   // IF ACELERATION STATE IS ACTIVE => SEND COMMAND TO GRADUALLY INCREASE MOTOR VELOCITY
         A     #Incremental_State;
         JCN   _100;

   // ANOLOG SIGNAL UNSCALING TO GENEREATE THE INCREMENTAL ACTION BASED ON A TIMER

         CALL  UNSCALE
         ( IN      := #Increment,
           HI_LIM  := #Max_Lim,
           LO_LIM  := #Low_Lim,
           BIPOLAR := FALSE,
           RET_VAL := #Ret_Val_Acel,
           OUT     := #Valve_Cmd
         );

   // SETTING THE MAX LIMIT
         L     #T_Increment;
         DTR;
         T     #Max_Lim;

   // MAPPING VAR FOR CONSULTING
         L     #Valve_Cmd;
         T     #PV;

   _100: NOP   0;

   // PERCENTAGE OF VALVE OPENED
         L     #Valve_Cmd;
         L     100;
         *I;
         T     "Tag_28";
         L     "Tag_28";
         L     27648;
         /I;
         DTR;
         RND;
         T     #"Vlv_Opened_%";


   // IF INCREMENTA STATE  = 1 AND NO TIMER.Q => SEND PULSE TO ACTIVATE TIMER
         A     #Incremental_State;
         AN    #Incremental_Timer.Q;
         =     #Pulse_Loop;


   // TIMER TO GENERATE THE INCREMENTAL VARIABLE
         CALL  #Incremental_Timer
         ( IN := #Pulse_Loop,
           PT := #T_Increment,
           Q  := ,
           ET := #Incremental_Timer.ET
         );


   // CONVERTIN THE ELAPSED TIME INTO REAL => TO ASIGN AS INPUT OF THE AO ACELERATION
         L     #Incremental_Timer.ET;
         DTR;
         T     #Increment;

   // MOTOR FEEDBACK
         L     #Valve_Cmd;
         L     0;
         >I;
         =     #Feedback;
END_REGION

REGION Network 2: CONDITIONS FOR EMERGENCY STOP BY OVERLOAD OR STOP BUTTON WHILE ACELERATING / /****************************** CLOSE MODE *****************************************/
   // IF MOTOR OVERLOAD OR STOP BUTTON AND ACELERATION => EMERGENCY STOP
         AN    #Vlv_Close_Cmd;
         FP    #FP_Stop;
         JCN   _108;
         L     0;
         T     #PV;
         T     #Increment;
         T     #Valve_Cmd;
         R     #Incremental_State;
   _108: NOP   0;
END_REGION

REGION Network 3: /******************************MANUAL MODE *****************************************/
   // MANUAL FULLY OPENED VALVE COMMAND
         A     #Manual;
         JCN   _2000;
         L     27648;
         T     #PV;
         L     100;
         T     #"Vlv_Opened_%";

   _2000:NOP   0;

   // MANUAL FULLY CLOSED VALVE COMMAND
         AN    #Manual;
         AN    #Incremental_State;
         JCN   _2001;
         L     0;
         T     #PV;

   _2001:NOP   0;
END_REGION
END_FUNCTION_BLOCK

(* ===== HMI "HMI_RT_1" =====
system functions are stored by id; their names below are inferred from use
connection "Conexión_1": ETHERNET, SIMATIC S7 300/400 MPI
connection "HMI_Conexión_1": ETHERNET, SIMATIC S7 300/400 MPI

HMI tags "Tabla de variables estándar"
   "TK101_FILLING_VLV_DB_Open_Valve_Cmd" : Bool = PLC TK101_FILLING_VLV_DB.Open_Valve_Cmd AT %DB3.DBX18.0, 1 s
   "Var_System_DB_Tk101_Level_%" : DInt = PLC Var_System_DB.Tk101.Level_% AT %DB1.DBD78, 100 ms
   "Var_System_DB_Tk102_Level_%" : DInt = PLC Var_System_DB.Tk102.Level_% AT %DB1.DBD128, 100 ms
   "Var_System_DB_Tk103_Level_%" : DInt = PLC Var_System_DB.Tk103.Level_% AT %DB1.DBD178, 100 ms
   "Var_System_DB_TK101_FILLING_VLV_Vlv_Cmd" : Bool = PLC Var_System_DB.TK101_FILLING_VLV.Vlv_Cmd AT %DB1.DBX106.0, 1 s
   "Var_System_DB_TK102_FILLING_VLV_Vlv_Cmd" : Bool = PLC Var_System_DB.TK102_FILLING_VLV.Vlv_Cmd AT %DB1.DBX156.0, 1 s
   "Var_System_DB_TK103_FILLING_VLV_Vlv_Cmd" : Bool = PLC Var_System_DB.TK103_FILLING_VLV.Vlv_Cmd AT %DB1.DBX206.0, 1 s
   "Var_System_DB_Weighing_Process_PV" : Real = PLC Var_System_DB.Weighing_Process.PV AT %DB1.DBD310, 1 s
   "Var_System_DB_Tk101_Vlv_Actuator_Cmd" : Int = PLC Var_System_DB.Tk101.Vlv_Actuator_Cmd AT %DB1.DBW66, 1 s
   "Var_System_DB_Tk101_High_Level_Alarm" : Bool = PLC Var_System_DB.Tk101.High_Level_Alarm AT %DB1.DBX62.5, 1 s
   "Var_System_DB_Tk101_Low_Level_Alarm" : Bool = PLC Var_System_DB.Tk101.Low_Level_Alarm AT %DB1.DBX62.4, 1 s
   "Var_System_DB_Tk102_Vlv_Actuator_Cmd" : Int = PLC Var_System_DB.Tk102.Vlv_Actuator_Cmd AT %DB1.DBW116, 1 s
   "Var_System_DB_Tk102_%_Vlv_Opened" : DInt = PLC Var_System_DB.Tk102.%_Vlv_Opened AT %DB1.DBD124, 1 s
   "Var_System_DB_Tk103_%_Vlv_Opened" : DInt = PLC Var_System_DB.Tk103.%_Vlv_Opened AT %DB1.DBD174, 1 s
   "Var_System_DB_Tk101_%_Vlv_Opened" : DInt = PLC Var_System_DB.Tk101.%_Vlv_Opened AT %DB1.DBD74, 1 s
   "Var_System_DB_Water_Valve_%_Vlv_Opened" : DInt = PLC Var_System_DB.Water_Valve.%_Vlv_Opened AT %DB1.DBD288, 1 s
   "Var_System_DB_Tk104_MIXER_Dis_Vlv_Cmd" : Bool = PLC Var_System_DB.Tk104_MIXER.Dis_Vlv_Cmd AT %DB1.DBX212.1, 1 s
   "HMI_VAR_Warnings" : Word = PLC HMI_VAR.Warnings AT %DB20.DBW22, 1 s
   "Var_System_DB_Tk101_Level_Liters" : Real = PLC Var_System_DB.Tk101.Level_Liters AT %DB1.DBD82, 1 s
   "Var_System_DB_TK101_FILLING_VLV_Vlv_Closed" : Bool = PLC Var_System_DB.TK101_FILLING_VLV.Vlv_Closed AT %DB1.DBX106.2, 1 s
   "Var_System_DB_TK101_FILLING_VLV_Vlv_Opened" : Bool = PLC Var_System_DB.TK101_FILLING_VLV.Vlv_Opened AT %DB1.DBX106.1, 1 s
   "Usuario" : WString[254], internal
   "Password" : WString[254], internal
   "HMI_VAR_Man_Valves_Filling_Vlv1" : Bool = PLC HMI_VAR.Man_Valves.Filling_Vlv1 AT %DB20.DBX24.0, 1 s
   "HMI_VAR_Man_Valves_Filling_Vlv2" : Bool = PLC HMI_VAR.Man_Valves.Filling_Vlv2 AT %DB20.DBX24.1, 1 s
   "HMI_VAR_Man_Valves_Filling_Vlv3" : Bool = PLC HMI_VAR.Man_Valves.Filling_Vlv3 AT %DB20.DBX24.2, 1 s
   "HMI_VAR_Man_Valves_Discharge_Vlv1" : Bool = PLC HMI_VAR.Man_Valves.Discharge_Vlv1 AT %DB20.DBX24.5, 1 s
   "HMI_VAR_Man_Valves_Discharge_Vlv2" : Bool = PLC HMI_VAR.Man_Valves.Discharge_Vlv2 AT %DB20.DBX24.6, 1 s
   "HMI_VAR_Man_Valves_Discharge_Vlv3" : Bool = PLC HMI_VAR.Man_Valves.Discharge_Vlv3 AT %DB20.DBX24.7, 1 s
   "HMI_VAR_Man_Valves_Scale_Vlv" : Bool = PLC HMI_VAR.Man_Valves.Scale_Vlv AT %DB20.DBX24.3, 1 s
   "HMI_VAR_Man_Valves_Mixer_Discharge_Vlv" : Bool = PLC HMI_VAR.Man_Valves.Mixer_Discharge_Vlv AT %DB20.DBX24.4, 1 s
   "HMI_VAR_Man_Valves_Water_Vlv" : Bool = PLC HMI_VAR.Man_Valves.Water_Vlv AT %DB20.DBX25.0, 1 s
   "HMI_VAR_Man_Valves_Sirupe_Vlv" : Bool = PLC HMI_VAR.Man_Valves.Sirupe_Vlv AT %DB20.DBX25.1, 1 s
   "HMI_VAR_Man_Motors_Conveyor" : Bool = PLC HMI_VAR.Man_Motors.Start_Conveyor AT %DB20.DBX26.0, 1 s
   "HMI_VAR_Man_Motors_Mixer" : Bool = PLC HMI_VAR.Man_Motors.Start_Mixer AT %DB20.DBX26.2, 1 s
   "Var_System_DB_TK102_FILLING_VLV_Vlv_Opened" : Bool = PLC Var_System_DB.TK102_FILLING_VLV.Vlv_Opened AT %DB1.DBX156.1, 1 s
   "Var_System_DB_TK102_FILLING_VLV_Vlv_Closed" : Bool = PLC Var_System_DB.TK102_FILLING_VLV.Vlv_Closed AT %DB1.DBX156.2, 1 s
   "Var_System_DB_TK103_FILLING_VLV_Vlv_Closed" : Bool = PLC Var_System_DB.TK103_FILLING_VLV.Vlv_Closed AT %DB1.DBX206.2, 1 s
   "Var_System_DB_TK103_FILLING_VLV_Vlv_Opened" : Bool = PLC Var_System_DB.TK103_FILLING_VLV.Vlv_Opened AT %DB1.DBX206.1, 1 s
   "Var_System_DB_Scale_Discharge_Vlv_Vlv_Opened" : Bool = PLC Var_System_DB.Scale_Discharge_Vlv.Vlv_Opened AT %DB1.DBX314.1, 1 s
   "Var_System_DB_Scale_Discharge_Vlv_Vlv_Closed" : Bool = PLC Var_System_DB.Scale_Discharge_Vlv.Vlv_Closed AT %DB1.DBX314.2, 1 s
   "Var_System_DB_Tk104_MIXER_Vlv_Closed" : Bool = PLC Var_System_DB.Tk104_MIXER.Vlv_Closed AT %DB1.DBX212.3, 1 s
   "Var_System_DB_Tk104_MIXER_Vlv_Opened" : Bool = PLC Var_System_DB.Tk104_MIXER.Vlv_Opened AT %DB1.DBX212.2, 1 s
   "Var_System_DB_Sirupe_Valve_%_Vlv_Opened" : DInt = PLC Var_System_DB.Sirupe_Valve.%_Vlv_Opened AT %DB1.DBD54, 1 s
   "Var_System_DB_Mixer_Motor_Feedback" : Bool = PLC Var_System_DB.Mixer_Motor.Feedback AT %DB1.DBX1.2, 1 s
   "Var_System_DB_Mixer_Motor_Led_Stopped" : Bool = PLC Var_System_DB.Mixer_Motor.Led_Stopped AT %DB1.DBX0.6, 1 s
   "Var_System_DB_Conveyor_Belt_M_Led_Stop" : Bool = PLC Var_System_DB.Conveyor_Belt.M_Led_Stop AT %DB1.DBX21.2, 1 s
   "Var_System_DB_Conveyor_Belt_M_Feedback" : Bool = PLC Var_System_DB.Conveyor_Belt.M_Feedback AT %DB1.DBX21.4, 1 s
   "Var_System_DB_Tk103_Vlv_Actuator_Cmd" : Int = PLC Var_System_DB.Tk103.Vlv_Actuator_Cmd AT %DB1.DBW166, 1 s
   "Var_System_DB_Sirupe_Valve_Vlv_Actuator_Cmd" : Int = PLC Var_System_DB.Sirupe_Valve.Vlv_Actuator_Cmd AT %DB1.DBW52, 1 s
   "Var_System_DB_Scale_Discharge_Vlv_Vlv_Cmd" : Bool = PLC Var_System_DB.Scale_Discharge_Vlv.Vlv_Cmd AT %DB1.DBX314.0, 1 s
   "Var_System_DB_Conveyor_Belt_M_Main" : Bool = PLC Var_System_DB.Conveyor_Belt.M_Main AT %DB1.DBX20.4, 1 s
   "Var_System_DB_Conveyor_Belt_M_Star" : Bool = PLC Var_System_DB.Conveyor_Belt.M_Star AT %DB1.DBX20.5, 1 s
   "Var_System_DB_Conveyor_Belt_M_Delta" : Bool = PLC Var_System_DB.Conveyor_Belt.M_Delta AT %DB1.DBX20.6, 1 s
   "HMI_VAR_Test_Recipe_Products{1}" : Real = PLC HMI_VAR.Test_Recipe.Products[1] AT %DB20.DBD2, 1 s
   "HMI_VAR_Test_Recipe_Products{2}" : Real = PLC HMI_VAR.Test_Recipe.Products[2] AT %DB20.DBD6, 1 s
   "HMI_VAR_Test_Recipe_Products{3}" : Real = PLC HMI_VAR.Test_Recipe.Products[3] AT %DB20.DBD10, 1 s
   "HMI_VAR_Test_Recipe_Flows{2}" : Real = PLC HMI_VAR.Test_Recipe.Flows[2] AT %DB20.DBD18, 1 s
   "HMI_VAR_Test_Recipe_Flows{1}" : Real = PLC HMI_VAR.Test_Recipe.Flows[1] AT %DB20.DBD14, 1 s
   "Var_System_DB_System_Generic_Start" : Bool = PLC Var_System_DB.System_Generic.Start AT %DB1.DBX12.2, 1 s
   "HMI_VAR_Conveyor_Container_Move" : Int = PLC HMI_VAR.Conveyor.Container_Move AT %DB20.DBW30, 100 ms
   "HMI_VAR_Mixer_Agitator_1" : Bool = PLC HMI_VAR.Mixer.Agitator_1 AT %DB20.DBX32.0, 100 ms
   "HMI_VAR_Mixer_Agitator_2" : Bool = PLC HMI_VAR.Mixer.Agitator_2 AT %DB20.DBX32.1, 100 ms
   "Var_System_DB_Tk104_MIXER_Level_%" : DInt = PLC Var_System_DB.Tk104_MIXER.Level_% AT %DB1.DBD234, 1 s
   "HMI_VAR_Conveyor_Belt" : Bool = PLC HMI_VAR.Conveyor.Belt AT %DB20.DBX28.0, 1 s
   "Var_System_DB_Conveyor_Belt_M_Led_Delta" : Bool = PLC Var_System_DB.Conveyor_Belt.M_Led_Delta AT %DB1.DBX21.1, 1 s
   "Var_System_DB_TK101_FILLING_VLV_Open_Vlv_Cmd" : Bool = PLC Var_System_DB.TK101_FILLING_VLV.Open_Vlv_Cmd AT %DB1.DBX106.4, 1 s
   "Var_System_DB_TK102_FILLING_VLV_Open_Vlv_Cmd" : Bool = PLC Var_System_DB.TK102_FILLING_VLV.Open_Vlv_Cmd AT %DB1.DBX156.4, 1 s
   "Var_System_DB_TK103_FILLING_VLV_Open_Vlv_Cmd" : Bool = PLC Var_System_DB.TK103_FILLING_VLV.Open_Vlv_Cmd AT %DB1.DBX206.4, 1 s
   "HMI_VAR_Recipe_Selection{1}" : Bool = PLC HMI_VAR.Recipe_Selection[1] AT %DB20.DBX0.0, 1 s
   "HMI_VAR_Recipe_Selection{2}" : Bool = PLC HMI_VAR.Recipe_Selection[2] AT %DB20.DBX0.1, 1 s
   "HMI_VAR_Recipe_Selection{3}" : Bool = PLC HMI_VAR.Recipe_Selection[3] AT %DB20.DBX0.2, 1 s
   "HMI_VAR_Reset_Selection" : Bool = PLC HMI_VAR.Reset_Selection AT %DB20.DBX34.5, 1 s
   "HMI_VAR_Start_Process" : Bool = PLC HMI_VAR.Start_Process AT %DB20.DBX34.4, 1 s
   "HMI_VAR_Recipe_Selection{4}" : Bool = PLC HMI_VAR.Recipe_Selection[4] AT %DB20.DBX0.3, 1 s
   "HMI_VAR_Enter_Selection" : Bool = PLC HMI_VAR.Enter_Selection AT %DB20.DBX34.3, 1 s
   "HMI_VAR_Auto/Manual" : Bool = PLC HMI_VAR.Auto/Manual AT %DB20.DBX34.2, 1 s
   "HMI_VAR_Act_System" : Bool = PLC HMI_VAR.Act_System AT %DB20.DBX34.0, 1 s
   "HMI_VAR_Stop_System" : Bool = PLC HMI_VAR.Stop_System AT %DB20.DBX34.1, 1 s
   "HMI_VAR_Man_Motors_Stop_Conveyor" : Bool = PLC HMI_VAR.Man_Motors.Stop_Conveyor AT %DB20.DBX26.1, 1 s
   "HMI_VAR_Man_Motors_Stop_Mixer" : Bool = PLC HMI_VAR.Man_Motors.Stop_Mixer AT %DB20.DBX26.3, 1 s
   "Var_System_DB_Scale_Discharge_Vlv_Open_Vlv_Cmd" : Bool = PLC Var_System_DB.Scale_Discharge_Vlv.Open_Vlv_Cmd AT %DB1.DBX314.5, 1 s
   "Scale_Dis_Vlv" : Bool = PLC Scale_Dis_Vlv AT %Q136.3, 1 s
   "Mixer_Dis_Vlv" : Bool = PLC Mixer_Dis_Vlv AT %Q136.4, 1 s

discrete alarms
   1: 'Overload Conveyor Motor', class Errors, trigger "HMI_VAR_Warnings" bit 0
      on Coming: function_f812520f('calvente.jaime@gmail.com', 'Fallo térmico del motor', 'El térmico ha saltado, por favor llamar técnico.', '')
   2: 'Overload Mixer Motor', class Errors, trigger "HMI_VAR_Warnings" bit 1
   3: 'Low level Tank 1', class Warnings, trigger "HMI_VAR_Warnings" bit 2
   4: 'High level Tank 1', class Warnings, trigger "HMI_VAR_Warnings" bit 3
   5: 'Low level Tank 2', class Warnings, trigger "HMI_VAR_Warnings" bit 4
   6: 'High level Tank 2', class Warnings, trigger "HMI_VAR_Warnings" bit 5
   7: 'Low level Tank 3', class Warnings, trigger "HMI_VAR_Warnings" bit 6
   8: 'High level Tank 3', class Warnings, trigger "HMI_VAR_Warnings" bit 7
   9: 'Emergency Stop', class Warnings, trigger "HMI_VAR_Warnings" bit 8

screen "GENERAL PROCESS" 1920x973, template "Plantilla_2"
   SymbolLibrary "Librería de símbolos_19" at 1370,493 size 306x261
   Bar "Barra_4" at 1410,521 size 225x182; MinimumValue 0; MaximumValue 100
      ProcessValue <- "Var_System_DB_Tk104_MIXER_Level_%"
   SymbolLibrary "Symbol library_2" at 1410,226 size 184x452
      Visibility <- "HMI_VAR_Mixer_Agitator_1"
   SymbolLibrary "Symbol library_3" at 1452,224 size 185x457
      Visibility <- "HMI_VAR_Mixer_Agitator_1"
   SymbolLibrary "Librería de símbolos_17" at 21,133 size 424x28
      Appearance <- "Var_System_DB_TK103_FILLING_VLV_Open_Vlv_Cmd"
   SymbolLibrary "Librería de símbolos_37" at 347,449 size 1097x344
   SymbolLibrary "Librería de símbolos_25" at 152,514 size 541x70
   SymbolLibrary "Librería de símbolos_11" at 131,271 size 190x182
   SymbolLibrary "Librería de símbolos_10" at 570,271 size 190x182
   SymbolLibrary "Librería de símbolos_12" at 348,271 size 190x182
   SymbolLibrary "Librería de símbolos_2" at 141,449 size 107x49
   SymbolLibrary "Librería de símbolos_3" at 357,448 size 108x50
   SymbolLibrary "Librería de símbolos_4" at 579,447 size 108x50
   SymbolLibrary "Librería de símbolos_5" at 203,494 size 45x26
   SymbolLibrary "Librería de símbolos_6" at 420,494 size 45x25
   SymbolLibrary "Librería de símbolos_7" at 642,492 size 45x27
   IOField "Campo ES_4" at 55,454 size 75x32; FormatPattern 999; Unit %
      ProcessValue <- "Var_System_DB_Tk101_%_Vlv_Opened"
   SymbolLibrary "Librería de símbolos_14" at 442,115 size 67x48
      Appearance <- "Var_System_DB_TK103_FILLING_VLV_Open_Vlv_Cmd"
   SymbolLibrary "Librería de símbolos_15" at 509,133 size 111x28
      Appearance <- "Var_System_DB_TK103_FILLING_VLV_Open_Vlv_Cmd"
   SymbolLibrary "Librería de símbolos_16" at 619,133 size 54x54
      Appearance <- "Var_System_DB_TK103_FILLING_VLV_Open_Vlv_Cmd"
   SymbolLibrary "Librería de símbolos_18" at 21,181 size 206x28
      Appearance <- "Var_System_DB_TK102_FILLING_VLV_Open_Vlv_Cmd"
   SymbolLibrary "Librería de símbolos_20" at 226,164 size 67x48
      Appearance <- "Var_System_DB_TK102_FILLING_VLV_Open_Vlv_Cmd"
   SymbolLibrary "Librería de símbolos_21" at 293,182 size 111x28
      Appearance <- "Var_System_DB_TK102_FILLING_VLV_Open_Vlv_Cmd"
   SymbolLibrary "Librería de símbolos_22" at 403,182 size 54x54
      Appearance <- "Var_System_DB_TK102_FILLING_VLV_Open_Vlv_Cmd"
   SymbolLibrary "Librería de símbolos_8" at 20,210 size 64x48
      Appearance <- "Var_System_DB_TK101_FILLING_VLV_Open_Vlv_Cmd"
   SymbolLibrary "Librería de símbolos_9" at 84,228 size 105x28
      Appearance <- "Var_System_DB_TK101_FILLING_VLV_Open_Vlv_Cmd"
   SymbolLibrary "Librería de símbolos_13" at 188,228 size 51x54
      Appearance <- "Var_System_DB_TK101_FILLING_VLV_Open_Vlv_Cmd"
   SymbolLibrary "Librería de símbolos_39" at 154,549 size 540x60
   SymbolLibrary "Librería de símbolos_40" at 356,607 size 135x42
   Bar "Barra_1" at 202,294 size 48x158; MinimumValue 0; MaximumValue 100
      ProcessValue <- "Var_System_DB_Tk101_Level_%"
   Bar "Barra_2" at 419,294 size 48x158; MinimumValue 0; MaximumValue 100
      ProcessValue <- "Var_System_DB_Tk102_Level_%"
   Bar "Barra_3" at 641,293 size 48x158; MinimumValue 0; MaximumValue 100
      ProcessValue <- "Var_System_DB_Tk103_Level_%"
   IOField "Campo ES_5" at 273,456 size 75x32; FormatPattern 999; Unit %
      ProcessValue <- "Var_System_DB_Tk102_%_Vlv_Opened"
   IOField "Campo ES_6" at 495,453 size 75x32; FormatPattern 999; Unit %
      ProcessValue <- "Var_System_DB_Tk103_%_Vlv_Opened"
   TextField "Campo de texto_7" at 541,18 size 890x81; Text 'PROCESS PLANT'
   IOField "Campo ES_3" at 154,521 size 141x49; FormatPattern 99999; Unit Kg
      ProcessValue <- "Var_System_DB_Weighing_Process_PV"
   SymbolLibrary "Librería de símbolos_26" at 1409,745 size 140x49
      Appearance <- "Var_System_DB_Tk104_MIXER_Dis_Vlv_Cmd"
   SymbolLibrary "Librería de símbolos_27" at 1491,702 size 71x47
   SymbolLibrary "Librería de símbolos_31" at 1801,450 size 104x97
   SymbolLibrary "Librería de símbolos_32" at 1676,517 size 130x24
   SymbolLibrary "Librería de símbolos_30" at 1801,556 size 104x96
   SymbolLibrary "Librería de símbolos_34" at 1674,622 size 131x24
   Group "Group_5" at 1514,793 size 184x43
   IOField "Campo ES_1" at 1699,484 size 92x32; FormatPattern 999; Unit %
      ProcessValue <- "Var_System_DB_Water_Valve_%_Vlv_Opened"
   SymbolLibrary "Symbol library_1" at 381,675 size 90x70
      DiagonalMovement <- "HMI_VAR_Conveyor_Container_Move"
   IOField "Campo ES_7" at 1582,240 size 132x55; FormatPattern 999; Unit %
      ProcessValue <- "Var_System_DB_Water_Valve_%_Vlv_Opened"
   IOField "Campo ES_2" at 1699,589 size 92x32; FormatPattern 999; Unit %
      ProcessValue <- "Var_System_DB_Sirupe_Valve_%_Vlv_Opened"
   TextField "Campo de texto_22" at 1332,232 size 230x66; Text 'AGITATOR VFD'
   SymbolLibrary "Symbol library_4" at 1472,321 size 119x118
   SymbolLibrary "Librería de símbolos_28" at 1514,793 size 49x43
   SymbolLibrary "Librería de símbolos_29" at 1561,815 size 137x21

screen "MENU" 1920x973, template "Plantilla_1"
   Button "Botón_1" at 125,225 size 1670x60; TextOff 'GENERAL PROCESS VISUALIZATION'
      on Press: ActivateScreen("GENERAL PROCESS", 0)
   Button "Botón_2" at 125,420 size 1670x60; TextOff 'RECIPE SELECTION'
      on Press: ActivateScreen("RECIPIES SELCTION", 0)
   Button "Botón_3" at 125,517 size 1670x60; TextOff 'AVISOS'
      on Press: ActivateScreen("WARNINGS", 0)
   Button "Botón_4" at 125,615 size 1670x60; TextOff 'GRAPHS'
      on Press: ActivateScreen("GRAPHS", 0)
   Button "Botón_5" at 125,715 size 1670x60; TextOff 'USERS'
      on Press: ActivateScreen("USERS", 0)
   TextField "Campo de texto_13" at 715,73 size 491x81; Text 'MAIN PLANT'
   Button "Botón_6" at 125,321 size 1670x60; TextOff 'MANUAL CONTROL PROCESS'; Authorization "Operación"
      on Press: ActivateScreen("MANUAL PROCESS", 0)

screen "TANKS" 1920x973, template "Plantilla_2"
   TextField "Campo de texto_13" at 387,9 size 1145x81; Text 'TANKS PROCESS VISUALIZATION'
   SymbolLibrary "Librería de símbolos_1" at 744,662 size 85x94
   IOField "Campo ES_3" at 1040,698 size 142x56; FormatPattern 999; Unit %
      ProcessValue <- "Var_System_DB_Tk102_Vlv_Actuator_Cmd"
   TextField "Campo de texto_5" at 951,635 size 232x39; Text 'DISCHARGE VLV 2'
   TextField "Campo de texto_6" at 861,155 size 232x40; Text 'TANK 2'
   TextField "Campo de texto_7" at 735,492 size 143x40; Text 'TANK LEVEL'
   TextField "Campo de texto_8" at 735,275 size 150x40; Text 'FILLING VLV 2'
   SymbolLibrary "Librería de símbolos_4" at 737,337 size 67x42
      Appearance <- "Var_System_DB_TK102_FILLING_VLV_Vlv_Cmd"
   IOField "Campo ES_4" at 735,551 size 138x38; FormatPattern 99; Unit %
      ProcessValue <- "Var_System_DB_Tk102_Level_%"
   SymbolLibrary "Librería de símbolos_5" at 1390,662 size 85x93
   IOField "Campo ES_5" at 1686,698 size 142x57; FormatPattern 999; Unit %
      ProcessValue <- "Var_System_DB_Tk103_Vlv_Actuator_Cmd"
   TextField "Campo de texto_9" at 1597,635 size 232x39; Text 'DISCHARGE VLV 3'
   TextField "Campo de texto_10" at 1507,155 size 232x40; Text 'TANK 3'
   TextField "Campo de texto_11" at 1381,492 size 143x40; Text 'TANK LEVEL'
   TextField "Campo de texto_12" at 1381,275 size 150x39; Text 'FILLING VLV 3'
   SymbolLibrary "Librería de símbolos_7" at 1384,337 size 67x42
      Appearance <- "Var_System_DB_TK103_FILLING_VLV_Vlv_Cmd"
   IOField "Campo ES_6" at 1382,551 size 138x38; FormatPattern 99; Unit %
      ProcessValue <- "Var_System_DB_Tk103_Level_%"
   Circle "Círculo_1" at 440,299 size 18x18
      Appearance <- "Var_System_DB_Tk101_High_Level_Alarm"
   Circle "Círculo_2" at 439,415 size 17x17
      Appearance <- "Var_System_DB_Tk101_Low_Level_Alarm"
   SymbolLibrary "Librería de símbolos_2" at 82,662 size 85x94
   IOField "Campo ES_1" at 378,698 size 142x56; FormatPattern 999; Unit %
      ProcessValue <- "Var_System_DB_Tk101_Vlv_Actuator_Cmd"
   TextField "Campo de texto_1" at 289,634 size 232x40; Text 'DISCHARGE VLV 1'
   TextField "Campo de texto_2" at 199,155 size 232x39; Text 'TANK 1'
   TextField "Campo de texto_3" at 73,492 size 143x40; Text 'TANK LEVEL'
   TextField "Campo de texto_4" at 73,275 size 150x39; Text 'FILLING VLV 1'
   SymbolLibrary "Librería de símbolos_14" at 76,334 size 67x42
      Appearance <- "Var_System_DB_TK103_FILLING_VLV_Vlv_Cmd"
   IOField "Campo ES_2" at 74,550 size 138x39; FormatPattern 99; Unit %
      ProcessValue <- "Var_System_DB_Tk101_Level_%"
   SymbolLibrary "Librería de símbolos_11" at 251,261 size 286x261
   Bar "Barra_1" at 351,294 size 85x145; MinimumValue 0; MaximumValue 100
      ProcessValue <- "Var_System_DB_Tk101_Level_%"
   SymbolLibrary "Librería de símbolos_3" at 913,262 size 286x259
   Bar "Barra_2" at 1013,294 size 85x145; MinimumValue 0; MaximumValue 100
      ProcessValue <- "Var_System_DB_Tk101_Level_%"
   SymbolLibrary "Librería de símbolos_6" at 1559,262 size 286x260
   Bar "Barra_3" at 1659,294 size 85x146; MinimumValue 0; MaximumValue 100
      ProcessValue <- "Var_System_DB_Tk103_Level_%"

screen "CONVEYOR" 1920x973, template "Plantilla_2"
   SymbolLibrary "Librería de símbolos_25" at 256,263 size 541x70
   SymbolLibrary "Librería de símbolos_39" at 258,318 size 540x60
   SymbolLibrary "Librería de símbolos_40" at 460,377 size 135x74
   SymbolLibrary "Librería de símbolos_1" at 280,612 size 120x120
   TextField "Campo de texto_5" at 543,612 size 232x39; Text 'DISCHARGE VLV'
   TextField "Campo de texto_6" at 415,152 size 232x40; Text 'SCALE'
   TextField "Campo de texto_7" at 251,463 size 175x44; Text 'WEIGHING'
   IOField "Campo ES_4" at 266,523 size 159x38; FormatPattern 999999; Unit kG
      ProcessValue <- "Var_System_DB_Weighing_Process_PV"
   TextField "Campo de texto_13" at 391,9 size 1141x81; Text 'WEIGHING PROCESS'
   SymbolLibrary "Librería de símbolos_2" at 1117,612 size 170x120
   TextField "Campo de texto_1" at 1267,153 size 228x40; Text 'CONVEYOR'
   SymbolLibrary "Symbol library_1" at 1117,333 size 524x120
   TextField "Campo de texto_4" at 1336,604 size 187x34; Text 'KM MAIN'
   TextField "Campo de texto_2" at 1337,651 size 187x34; Text 'KM STAR'
   TextField "Campo de texto_3" at 1337,700 size 187x34; Text 'KM DELTA'
   TextField "Campo de texto_10" at 601,670 size 164x57; Text 'CLOSED'
      Visibility <- "Var_System_DB_Scale_Discharge_Vlv_Vlv_Cmd"
   TextField "Campo de texto_11" at 601,669 size 164x58; Text 'OPENED'
      Visibility <- "Var_System_DB_Scale_Discharge_Vlv_Vlv_Cmd"
   TextField "Campo de texto_18" at 1561,605 size 83x33; Text 'ON'
      Visibility <- "Var_System_DB_Conveyor_Belt_M_Main"
   TextField "Campo de texto_19" at 1561,605 size 83x33; Text 'OFF'
      Visibility <- "Var_System_DB_Conveyor_Belt_M_Main"
   TextField "Campo de texto_8" at 1561,651 size 83x33; Text 'ON'
      Visibility <- "Var_System_DB_Conveyor_Belt_M_Star"
   TextField "Campo de texto_9" at 1561,651 size 83x33; Text 'OFF'
      Visibility <- "Var_System_DB_Conveyor_Belt_M_Star"
   TextField "Campo de texto_12" at 1561,697 size 83x33; Text 'ON'
      Visibility <- "Var_System_DB_Conveyor_Belt_M_Led_Delta"
   TextField "Campo de texto_14" at 1561,697 size 83x33; Text 'OFF'
      Visibility <- "Var_System_DB_Conveyor_Belt_M_Led_Delta"

screen "MIXER" 1920x973, template "Plantilla_2"
   SymbolLibrary "Librería de símbolos_2" at 412,342 size 367x332
   Bar "Barra_1" at 504,377 size 188x223; MinimumValue 0; MaximumValue 100
      ProcessValue <- "Var_System_DB_Tk103_Level_%"
   SymbolLibrary "Librería de símbolos_3" at 1253,318 size 137x74
   IOField "Campo ES_1" at 1405,340 size 182x53; FormatPattern 999; Unit %
      ProcessValue <- "Var_System_DB_Water_Valve_%_Vlv_Opened"
   IOField "Campo ES_2" at 1416,482 size 171x49; FormatPattern 999; Unit %
      ProcessValue <- "Var_System_DB_Sirupe_Valve_%_Vlv_Opened"
   SymbolLibrary "Librería de símbolos_6" at 998,164 size 261x95
   Button "Botón_14" at 407,184 size 489x65; TextOff 'MIXER MOTOR'
      on Press: function_b14e0dd5("HMI_VAR_Man_Motors_Mixer", 0)
   TextField "Campo de texto_20" at 1329,191 size 185x53; Text 'OFF'
      Visibility <- "Var_System_DB_Mixer_Motor_Feedback"
   TextField "Campo de texto_21" at 1329,191 size 185x53; Text 'ON'
      Visibility <- "Var_System_DB_Mixer_Motor_Feedback"
   IOField "Campo ES_10" at 639,727 size 166x52; FormatPattern 999; Unit %
      ProcessValue <- "Var_System_DB_Tk101_Level_%"
   TextField "Campo de texto_23" at 374,725 size 245x54; Text 'TK4 LEVEL'
   Button "Botón_16" at 880,342 size 347x47; TextOff 'WATER VALVE'
      on Press: function_b14e0dd5("HMI_VAR_Man_Valves_Water_Vlv", 0)
   SymbolLibrary "Librería de símbolos_7" at 1252,457 size 135x77
   Button "Botón_17" at 878,482 size 347x46; TextOff 'SIRUPE VALVE'
      on Press: function_b14e0dd5("HMI_VAR_Man_Valves_Sirupe_Vlv", 0)
   Button "Botón_18" at 872,616 size 346x48; TextOff 'DISCHARGE VALVE'
      on Press: function_b14e0dd5("HMI_VAR_Man_Valves_Mixer_Discharge_Vlv", 0)
   SymbolLibrary "Librería de símbolos_4" at 1272,592 size 90x80
      Appearance <- "Var_System_DB_Tk104_MIXER_Dis_Vlv_Cmd"
   TextField "Campo de texto_24" at 1391,608 size 186x55; Text 'OPENED'
      Visibility <- "Var_System_DB_Tk104_MIXER_Dis_Vlv_Cmd"
   TextField "Campo de texto_25" at 1392,608 size 186x55; Text 'CLOSED'
      Visibility <- "Var_System_DB_Tk104_MIXER_Dis_Vlv_Cmd"
   TextField "Campo de texto_7" at 388,17 size 1145x81; Text 'MIXER STATION'

Template "Plantilla_2" 1920x973
   Button "Botón_1" at 15,854 size 132x106; TextOff 'Text'; PictureOff "Home"
      on Press: ActivateScreen("MENU", 0)
   Button "Botón_2" at 589,855 size 132x106; TextOff 'TANKS'; PictureOff "Home"; Authorization "Operación"
      on Press: ActivateScreen("TANKS", 0)
   Button "Botón_3" at 785,855 size 132x106; TextOff 'CONVEYOR'; PictureOff "Home"; Authorization "Operación"
      on Press: ActivateScreen("CONVEYOR", 0)
   Button "Botón_4" at 981,855 size 132x106; TextOff 'MIXER'; PictureOff "Home"; Authorization "Operación"
      on Press: ActivateScreen("MIXER", 0)
   Button "Botón_7" at 1359,855 size 262x106; TextOff 'START'; PictureOff "Home"; Authorization "Administración de usuarios"
      on Press: function_b14e0dd5("HMI_VAR_Act_System", 0)
   Button "Botón_8" at 1647,855 size 263x106; TextOff 'STOP'; PictureOff "Home"; Authorization "Administración de usuarios"
      on Press: function_b14e0dd5("HMI_VAR_Stop_System", 0)
   Button "Botón_5" at 205,855 size 132x106; TextOff 'GENERAL'; PictureOff "Home"; Authorization "Operación"
      on Press: ActivateScreen("GENERAL PROCESS", 0)
   Button "Botón_10" at 398,854 size 132x106; TextOff 'MANUAL'; PictureOff "Home"; Authorization "Operación"
      on Press: ActivateScreen("MANUAL PROCESS", 0)

screen "RECIPIES SELCTION" 1920x973, template "Plantilla_2"
   Button "Botón_1" at 125,188 size 1670x92; TextOff 'RECIPE 1'
      on Press: function_b14e0dd5("HMI_VAR_Recipe_Selection{1}", 0)
   Button "Botón_2" at 125,325 size 1670x92; TextOff 'RECIPE 2'
      on Press: function_b14e0dd5("HMI_VAR_Recipe_Selection{2}", 0)
   Button "Botón_3" at 125,466 size 1670x92; TextOff 'RECIPE 3'
      on Press: function_b14e0dd5("HMI_VAR_Recipe_Selection{3}", 0)
   Button "Botón_4" at 125,593 size 1670x92; TextOff 'TEST RECIPE'; Authorization "Administración de usuarios"
      on Press: ActivateScreen("RECIPE TEST", 0); function_b14e0dd5("HMI_VAR_Recipe_Selection{4}", 0)
   TextField "Campo de texto_13" at 592,73 size 737x81; Text 'RECIPE SELECTION'
   Button "Button_1" at 352,725 size 327x67; TextOff 'RESET SELECTION'
      on Press: function_b14e0dd5("HMI_VAR_Reset_Selection", 0)
   Button "Button_2" at 1290,727 size 327x67; TextOff 'START PROCESS'
      on Press: function_b14e0dd5("HMI_VAR_Enter_Selection", 0)

screen "RECIPE TEST" 1920x973, template "Plantilla_2"
   TextField "Campo de texto_7" at 552,42 size 816x82; Text 'TEST RECIPE'
   Button "Botón_1" at 163,156 size 384x50; TextOff 'PRODUCT A'
      on Press: ActivateScreen("GENERAL PROCESS", 0)
   IOField "I/O field_1" at 1487,151 size 245x52; FormatPattern 999999; Unit Kg
      ProcessValue <- "HMI_VAR_Test_Recipe_Products{1}"
   Button "Botón_2" at 163,263 size 384x48; TextOff 'PRODUCT B'
      on Press: ActivateScreen("GENERAL PROCESS", 0)
   IOField "I/O field_2" at 1487,259 size 245x50; FormatPattern 999999; Unit Kg
      ProcessValue <- "HMI_VAR_Test_Recipe_Products{2}"
   Button "Botón_3" at 163,366 size 384x49; TextOff 'PRODUCT C'
      on Press: ActivateScreen("GENERAL PROCESS", 0)
   IOField "I/O field_3" at 1487,362 size 245x51; FormatPattern 999999; Unit Kg
      ProcessValue <- "HMI_VAR_Test_Recipe_Products{3}"
   Button "Botón_4" at 163,466 size 384x49; TextOff 'WATER FLOW'
      on Press: ActivateScreen("GENERAL PROCESS", 0)
   IOField "I/O field_4" at 1487,462 size 245x50; FormatPattern 99; Unit L/S
      ProcessValue <- "HMI_VAR_Test_Recipe_Flows{1}"
   Button "Botón_5" at 163,567 size 384x49; TextOff 'SYRUPE FLOW'
      on Press: ActivateScreen("GENERAL PROCESS", 0)
   IOField "I/O field_5" at 1487,562 size 245x52; FormatPattern 99; Unit L/S
      ProcessValue <- "HMI_VAR_Test_Recipe_Flows{2}"
   Button "Button_1" at 723,711 size 474x96; TextOff 'START PROCESS'
      on Press: function_b14e0dd5("HMI_VAR_Enter_Selection", 0)

screen "GRAPHS" 1920x973, template "Plantilla_2"
   TrendView "Visor de curvas_1" at 195,171 size 1504x590

screen "WARNINGS" 1920x973, template "Plantilla_2"
   AlarmView "Visor de avisos_1" at 324,116 size 1273x311
   AlarmView "Visor de avisos_2" at 324,510 size 1273x319
   TextField "Campo de texto_7" at 515,13 size 890x81; Text 'WARININGS'

screen "MANUAL PROCESS" 1920x973, template "Plantilla_2"
   SymbolLibrary "Librería de símbolos_25" at 725,563 size 541x58
   SymbolLibrary "Librería de símbolos_11" at 701,215 size 170x167
   SymbolLibrary "Librería de símbolos_10" at 1121,215 size 170x167
   SymbolLibrary "Librería de símbolos_12" at 907,215 size 170x167
   SymbolLibrary "Librería de símbolos_14" at 395,206 size 74x45
      Appearance <- "Var_System_DB_TK103_FILLING_VLV_Vlv_Cmd"
   SymbolLibrary "Librería de símbolos_39" at 726,607 size 540x48
   SymbolLibrary "Librería de símbolos_40" at 928,654 size 135x30
   Bar "Barra_1" at 771,238 size 28x143; MinimumValue 0; MaximumValue 100
      ProcessValue <- "Var_System_DB_Tk101_Level_%"
   Bar "Barra_2" at 978,239 size 28x143; MinimumValue 0; MaximumValue 100
      ProcessValue <- "Var_System_DB_Tk102_Level_%"
   Bar "Barra_3" at 1192,238 size 28x143; MinimumValue 0; MaximumValue 100
      ProcessValue <- "Var_System_DB_Tk103_Level_%"
   TextField "Campo de texto_1" at 513,212 size 83x33; Text 'OPENED'
      Visibility <- "Var_System_DB_TK101_FILLING_VLV_Open_Vlv_Cmd"
   TextField "Campo de texto_2" at 513,212 size 83x33; Text 'CLOSED'
      Visibility <- "Var_System_DB_TK101_FILLING_VLV_Open_Vlv_Cmd"
   Button "Botón_15" at 72,211 size 285x40; TextOff 'MANUAL VALVE 1'
      on Press: function_b14e0dd5("HMI_VAR_Man_Valves_Filling_Vlv1", 0)
   SymbolLibrary "Librería de símbolos_8" at 394,294 size 74x45
      Appearance <- "Var_System_DB_TK103_FILLING_VLV_Vlv_Cmd"
   TextField "Campo de texto_3" at 508,303 size 83x33; Text 'OPENED'
      Visibility <- "Var_System_DB_TK102_FILLING_VLV_Open_Vlv_Cmd"
   TextField "Campo de texto_4" at 508,303 size 83x33; Text 'CLOSED'
      Visibility <- "Var_System_DB_TK102_FILLING_VLV_Open_Vlv_Cmd"
   Button "Botón_9" at 71,299 size 285x40; TextOff 'MANUAL VALVE 2'
      on Press: function_b14e0dd5("HMI_VAR_Man_Valves_Filling_Vlv2", 0)
   SymbolLibrary "Librería de símbolos_9" at 395,379 size 74x45
      Appearance <- "Var_System_DB_TK103_FILLING_VLV_Vlv_Cmd"
   TextField "Campo de texto_5" at 509,388 size 83x33; Text 'OPENED'
      Visibility <- "Var_System_DB_TK103_FILLING_VLV_Open_Vlv_Cmd"
   TextField "Campo de texto_6" at 509,388 size 83x33; Text 'CLOSED'
      Visibility <- "Var_System_DB_TK103_FILLING_VLV_Open_Vlv_Cmd"
   Button "Botón_10" at 72,384 size 285x40; TextOff 'MANUAL VALVE 3'
      on Press: function_b14e0dd5("HMI_VAR_Man_Valves_Filling_Vlv3", 0)
   TextField "Campo de texto_13" at 186,139 size 310x42; Text 'FILLING VALVES'
   TextField "Campo de texto_7" at 388,17 size 1145x81; Text 'MANUAL PROCESS'
   Button "Botón_5" at 72,560 size 285x40; TextOff 'MANUAL VALVE 1'
      on Press: function_b14e0dd5("HMI_VAR_Man_Valves_Discharge_Vlv1", 0)
   Button "Botón_11" at 71,648 size 285x40; TextOff 'MANUAL VALVE 2'
      on Press: function_b14e0dd5("HMI_VAR_Man_Valves_Discharge_Vlv2", 0)
   Button "Botón_12" at 72,733 size 285x40; TextOff 'MANUAL VALVE 3'
      on Press: function_b14e0dd5("HMI_VAR_Man_Valves_Discharge_Vlv3", 0)
   TextField "Campo de texto_15" at 148,491 size 369x38; Text 'DISCHARGE VALVES'
   SymbolLibrary "Librería de símbolos_2" at 412,546 size 49x64
   IOField "Campo ES_4" at 516,568 size 75x32; FormatPattern 999; Unit %
      ProcessValue <- "Var_System_DB_Tk101_%_Vlv_Opened"
   IOField "Campo ES_5" at 518,648 size 75x32; FormatPattern 999; Unit %
      ProcessValue <- "Var_System_DB_Tk102_%_Vlv_Opened"
   IOField "Campo ES_6" at 517,739 size 75x32; FormatPattern 999; Unit %
      ProcessValue <- "Var_System_DB_Tk103_%_Vlv_Opened"
   SymbolLibrary "Librería de símbolos_3" at 413,634 size 49x64
   SymbolLibrary "Librería de símbolos_4" at 414,720 size 49x64
   TextField "Campo de texto_8" at 839,140 size 310x42; Text 'TANKS LEVELS'
   TextField "Campo de texto_9" at 845,490 size 310x42; Text 'SCALE'
   IOField "Campo ES_3" at 725,565 size 144x46; FormatPattern 99999; Unit Kg
      ProcessValue <- "Var_System_DB_Weighing_Process_PV"
   Button "Botón_13" at 725,743 size 240x40; TextOff 'MANUAL SCALE VLV'
      on Press: function_b14e0dd5("HMI_VAR_Man_Valves_Scale_Vlv", 0)
   SymbolLibrary "Librería de símbolos_5" at 1021,738 size 74x45
      Appearance <- "Var_System_DB_TK103_FILLING_VLV_Vlv_Cmd"
   TextField "Campo de texto_10" at 1142,748 size 83x33; Text 'CLOSED'
      Visibility <- "Var_System_DB_Scale_Discharge_Vlv_Open_Vlv_Cmd"
   TextField "Campo de texto_11" at 1142,748 size 83x33; Text 'OPENED'
      Visibility <- "Scale_Dis_Vlv"
   SymbolLibrary "Librería de símbolos_1" at 1621,209 size 117x58
   IOField "Campo ES_7" at 809,413 size 75x32; FormatPattern 999; Unit %
      ProcessValue <- "Var_System_DB_Tk101_Level_%"
   IOField "Campo ES_8" at 1017,413 size 75x32; FormatPattern 999; Unit %
      ProcessValue <- "Var_System_DB_Tk102_Level_%"
   IOField "Campo ES_9" at 1228,413 size 75x32; FormatPattern 999; Unit %
      ProcessValue <- "Var_System_DB_Tk103_Level_%"
   TextField "Campo de texto_12" at 691,412 size 110x33; Text 'TK1 LEVEL'
   TextField "Campo de texto_14" at 899,412 size 110x33; Text 'TK2 LEVEL'
   TextField "Campo de texto_16" at 1105,411 size 110x33; Text 'TK3 LEVEL'
   TextField "Campo de texto_17" at 1469,140 size 310x42; Text 'CONVEYOR MOTOR'
   Button "Botón_1" at 1356,221 size 96x40; TextOff 'START'
      on Press: function_b14e0dd5("HMI_VAR_Man_Motors_Conveyor", 0)
   TextField "Campo de texto_18" at 1771,222 size 83x33; Text 'ON'
      Visibility <- "Var_System_DB_Conveyor_Belt_M_Main"
   TextField "Campo de texto_19" at 1771,222 size 83x33; Text 'OFF'
      Visibility <- "Var_System_DB_Conveyor_Belt_M_Main"
   Button "Botón_4" at 1459,221 size 96x40; TextOff 'STOP'
      on Press: function_b14e0dd5("HMI_VAR_Man_Motors_Stop_Conveyor", 0)
   SymbolLibrary "Librería de símbolos_19" at 1361,516 size 166x203
   SymbolLibrary "Librería de símbolos_31" at 1741,502 size 61x45
   IOField "Campo ES_1" at 1809,515 size 82x33; FormatPattern 999; Unit %
      ProcessValue <- "Var_System_DB_Water_Valve_%_Vlv_Opened"
   IOField "Campo ES_2" at 1814,601 size 77x31; FormatPattern 999; Unit %
      ProcessValue <- "Var_System_DB_Sirupe_Valve_%_Vlv_Opened"
   SymbolLibrary "Librería de símbolos_6" at 1626,408 size 117x58
   TextField "Campo de texto_20" at 1775,424 size 83x33; Text 'OFF'
      Visibility <- "Var_System_DB_Mixer_Motor_Feedback"
   TextField "Campo de texto_21" at 1775,424 size 83x33; Text 'ON'
      Visibility <- "Var_System_DB_Mixer_Motor_Feedback"
   TextField "Campo de texto_22" at 1474,338 size 310x42; Text 'MIXER STATION'
   IOField "Campo ES_10" at 1464,751 size 75x32; FormatPattern 999; Unit %
      ProcessValue <- "Var_System_DB_Tk101_Level_%"
   TextField "Campo de texto_23" at 1345,750 size 110x33; Text 'TK4 LEVEL'
   Button "Botón_16" at 1573,516 size 156x29; TextOff 'WATER VALVE'
      on Press: function_b14e0dd5("HMI_VAR_Man_Valves_Water_Vlv", 0)
   SymbolLibrary "Librería de símbolos_7" at 1740,587 size 61x45
   Button "Botón_17" at 1572,601 size 156x29; TextOff 'SIRUPE VALVE'
      on Press: function_b14e0dd5("HMI_VAR_Man_Valves_Sirupe_Vlv", 0)
   Button "Botón_18" at 1569,684 size 156x29; TextOff 'DISCHARGE VLV'
      on Press: function_b14e0dd5("HMI_VAR_Man_Valves_Mixer_Discharge_Vlv", 0)
   SymbolLibrary "Librería de símbolos_26" at 1749,669 size 41x49
      Appearance <- "Var_System_DB_Tk104_MIXER_Dis_Vlv_Cmd"
   TextField "Campo de texto_24" at 1803,679 size 83x33; Text 'OPENED'
      Visibility <- "Mixer_Dis_Vlv"
   TextField "Campo de texto_25" at 1803,679 size 83x33; Text 'CLOSED'
      Visibility <- "Mixer_Dis_Vlv"
   Button "Botón_6" at 1356,419 size 96x40; TextOff 'START'
      on Press: function_b14e0dd5("HMI_VAR_Man_Motors_Mixer", 0)
   Button "Botón_7" at 1459,420 size 96x40; TextOff 'STOP'
      on Press: function_b14e0dd5("HMI_VAR_Man_Motors_Stop_Mixer", 0)
   Bar "Barra_4" at 1394,538 size 102x134; MinimumValue 0; MaximumValue 100
      ProcessValue <- "Var_System_DB_Tk104_MIXER_Level_%"

screen "PORTAL" 1920x973
   GraphicView "Graphic view_1" at 0,4 size 1918x966; Picture "depositphotos_88642944-stock-illustration-industrial-plant-factory-site"
   Button "Botón_1" at 1239,792 size 610x120; TextOff 'GO TO PROCESS'; Authorization "Operación"
      on Press: ActivateScreen("MAN/AUTO", 0)

screen "MAN/AUTO" 1920x973, template "Plantilla_1"
   Button "Button_1" at 400,339 size 381x171; TextOff 'AUTO'
      on Press: ResetBit("HMI_VAR_Auto/Manual"); ActivateScreen("GENERAL PROCESS", 0)
   Button "Button_2" at 1098,343 size 381x171; TextOff 'MANUAL'
      on Press: SetBit("HMI_VAR_Auto/Manual"); ActivateScreen("MANUAL PROCESS", 0)
   TextField "Campo de texto_13" at 437,47 size 1047x107; Text 'RECIPE SELECTION'
*)